
                                #statStateMQTTinternal := #IDLE;
                            END_IF;
                        ELSIF #instTcpSend.ERROR
                        THEN
                            #statusID := #MQTT_PUBLISH;
                            #instTcpSend.REQ := false;
                            #statStateMQTT := #MQTT_ERROR;
                            #status := #instTcpSend.STATUS;
                        END_IF;
                    #MQTT_PUBACK:
                        IF #statNewDataRcv THEN
                            IF ((#statRcvBuffer[1] AND b#16#f0) = #MQTT_MSG_TYPE_PUBACK)
                                OR
                                ((#statRcvBuffer[1] AND b#16#f0) = INT_TO_WORD(#MQTT_MSG_TYPE_PUBREC))
                            THEN
                                IF
                                    (#statRcvBuffer[3] = #statPacketIDAck.%B1)
                                    AND
                                    (#statRcvBuffer[4] = #statPacketIDAck.%B0)
                                THEN
                                    IF (#mqttParam.publishFlag.qualityOfService = 1)
                                    THEN
                                        //QoS = 1; finish here
                                        #statStateMQTTinternal := #MQTT_IDLE;
                                        #published := true;
                                        #busy := false;
                                        #statNewDataRcv := false;
                                        //Re-Activate Kepp Alive Timer
                                        IF NOT #statKeepAliveOff
                                        THEN
                                            #statTriggerKeepAlive := true;
                                        END_IF;

                                        #statStateMQTTinternal := #IDLE;
                                    ELSE
                                        #statStateMQTTinternal := #MQTT_PUBREL;
                                    END_IF;
                                ELSE
                                    #statNewDataRcv := false;
                                END_IF;
                            ELSE
                                #statStateMQTT := #MQTT_ERROR;
                                #statusID := #MQTT_PUBACK;
                            END_IF;
                        END_IF;
                    #MQTT_PUBREL:
                        //fixed Header
                        #statSendBuffer[1] := 16#62;
                        #statSendBuffer[2] := 2;
                        //Variable Header
                        #statSendBuffer[3] := #statPacketID.%B1;
                        #statSendBuffer[4] := #statPacketID.%B0;
                        #instTcpSend.LEN := INT_TO_UDINT(4);
                        #instTcpSend.REQ := true;

                        IF ((#instTcpSend.DONE)
                            AND (#instTcpSend.BUSY = 0))
                        THEN
                            #instTcpSend.REQ := false;
                            #statPacketIDAck := #statPacketID;
                            #statStateMQTTinternal := #MQTT_PUBCOMP;

                        ELSIF #instTcpSend.ERROR
                        THEN
                            #statusID := #MQTT_PUBREL;
                            #instTcpSend.REQ := false;
                            #statStateMQTT := #MQTT_ERROR;
                            #status := #instTcpSend.STATUS;
                        END_IF;
                    #MQTT_PUBCOMP:
                        IF #statNewDataRcv THEN
                            IF ((#statRcvBuffer[1] AND b#16#f0) = #MQTT_MSG_TYPE_PUBCOM)
                            THEN
                                IF
                                    (#statRcvBuffer[3] = #statPacketIDAck.%B1)
                                    AND
                                    (#statRcvBuffer[4] = #statPacketIDAck.%B0)
                                THEN
                                    //QoS = 2; finish here
                                    #statStateMQTTinternal := #MQTT_IDLE;
                                    #published := true;
                                    #busy := false;
                                    #statNewDataRcv := false;
                                    //Re-Activate Kepp Alive Timer
                                    IF NOT #statKeepAliveOff
                                    THEN
                                        #statTriggerKeepAlive := true;
                                    END_IF;

                                    #statStateMQTTinternal := #IDLE;
                                ELSE
                                    #statStateMQTT := #MQTT_ERROR;
                                    #statusID := #MQTT_PUBCOMP;
                                END_IF;
                            END_IF;
                        END_IF;
                    #MQTT_PING:

                        #busy := true;
                        //Build fixed Header
                        //Message Type
                        #statSendBuffer[1] := INT_TO_BYTE(#MQTT_MSG_TYPE_PING);
                        //Remaining Lenght (must be O)
                        #statSendBuffer[2] := 0;
                        #instTcpSend.REQ := true;
                        #instTcpSend.LEN := 2;

                        IF ((#instTcpSend.DONE)
                            AND (#instTcpSend.BUSY = 0))
                        THEN
                            #instTcpSend.REQ := false;
                            #statStateMQTTinternal := #MQTT_PINGRESP;
                        ELSIF #instTcpSend.ERROR
                        THEN
                            #statusID := #MQTT_PING;
                            #instTcpSend.REQ := false;
                            #statStateMQTT := #MQTT_ERROR;
                            #status := #instTcpSend.STATUS;
                        END_IF;
                    #MQTT_PINGRESP:
                        IF #statNewDataRcv
                        THEN
                            IF ((#statRcvBuffer[1] AND b#16#f0) = #MQTT_MSG_TYPE_PINGRESP)
                            THEN
                                #busy := false;
                                #statNewDataRcv := false;
                                #statTriggerKeepAlive := true;
                                #statStateMQTTinternal := #IDLE;
                            END_IF;
                        ELSE
                            #statNewDataRcv := false;
                        END_IF;

                END_CASE;
           #MQTT_DISCONNECT:
           #busy := 0;
           //Build fixed Header
           //Message Type
           #statSendBuffer[1] := INT_TO_BYTE(#MQTT_MSG_TYPE_DISCONNECT);
           //Remaining Lenght (must be O)
           #statSendBuffer[2] := 0;
           #instTcpSend.REQ := true;
           #instTcpSend.LEN := 2;

           IF ((#instTcpSend.DONE)
               AND (#instTcpSend.BUSY = 0))
           THEN
               IF NOT #enable THEN
                   #statStateTCP := #TCP_DISCONNECT;
               END_IF;
               #instTcpSend.REQ := false;
               #statStateMQTT := #MQTT_DISCONNECTED;
               #statStateMQTTinternal := #IDLE;
           ELSIF #instTcpSend.ERROR
           THEN
               IF NOT #enable THEN
                   #statStateTCP := #TCP_DISCONNECT;
               END_IF;
               #statusID := #MQTT_DISCONNECT;
               #instTcpSend.REQ := false;
               #statStateMQTT := #MQTT_ERROR;
               #status := #instTcpSend.STATUS;
           END_IF;
               #MQTT_ERROR:

               REGION Errorhandling MQTT
                   #error := true;
                   #busy := false;
                   #statStateMQTTinternal := #IDLE;
                   #statTriggerKeepAlive := 0;
                   #statKeepAliveOff := false;
                 CASE #statusID OF
                     #MQTT_CONNECT_FLAG_CHECK:
                         #mqttEstablished := false;
                         #statStateMQTT := #MQTT_DISCONNECTED;
                         ;
                     #MQTT_CONNECT:
                         #mqttEstablished := false;
                         #status := #instTcpSend.STATUS;   ;
                         #statStateMQTT := #MQTT_DISCONNECTED;
                       #MQTT_CONNACK:
                           #mqttEstablished := false;
                           #status := #statRcvBuffer[4];
                           #statStateMQTT := #MQTT_DISCONNECTED;
                       #MQTT_PUBLISH:
                               #published := false;
                               #statStateMQTT := #MQTT_CONNECTED;
                               #MQTT_PUBACK,#MQTT_PUBCOMP,#MQTT_PUBREL:
                           #published := false;
                           #status :=#MQTT_ERROR_PACKETID;
                           #statStateMQTT := #MQTT_CONNECTED;
                       #MQTT_PINGRESP:;
                           #MQTT_PING:;
                       #MQTT_DISCONNECT:
                           #mqttEstablished := false;
                          ;
                       ELSE
                           ;
                   END_CASE;
              END_REGION
               ;



       END_CASE
       ;
END_FUNCTION_BLOCK

// folder: NodeRed

FUNCTION "FC_saveMotorDatatoDB" : Void   // FC13, LAD
{ S7_Optimized_Access := 'TRUE' }
VERSION : 0.1
BEGIN

REGION Network 1: M1
   // -temepratura
   // -status POS1
   // -status POS2
   // -isINerror
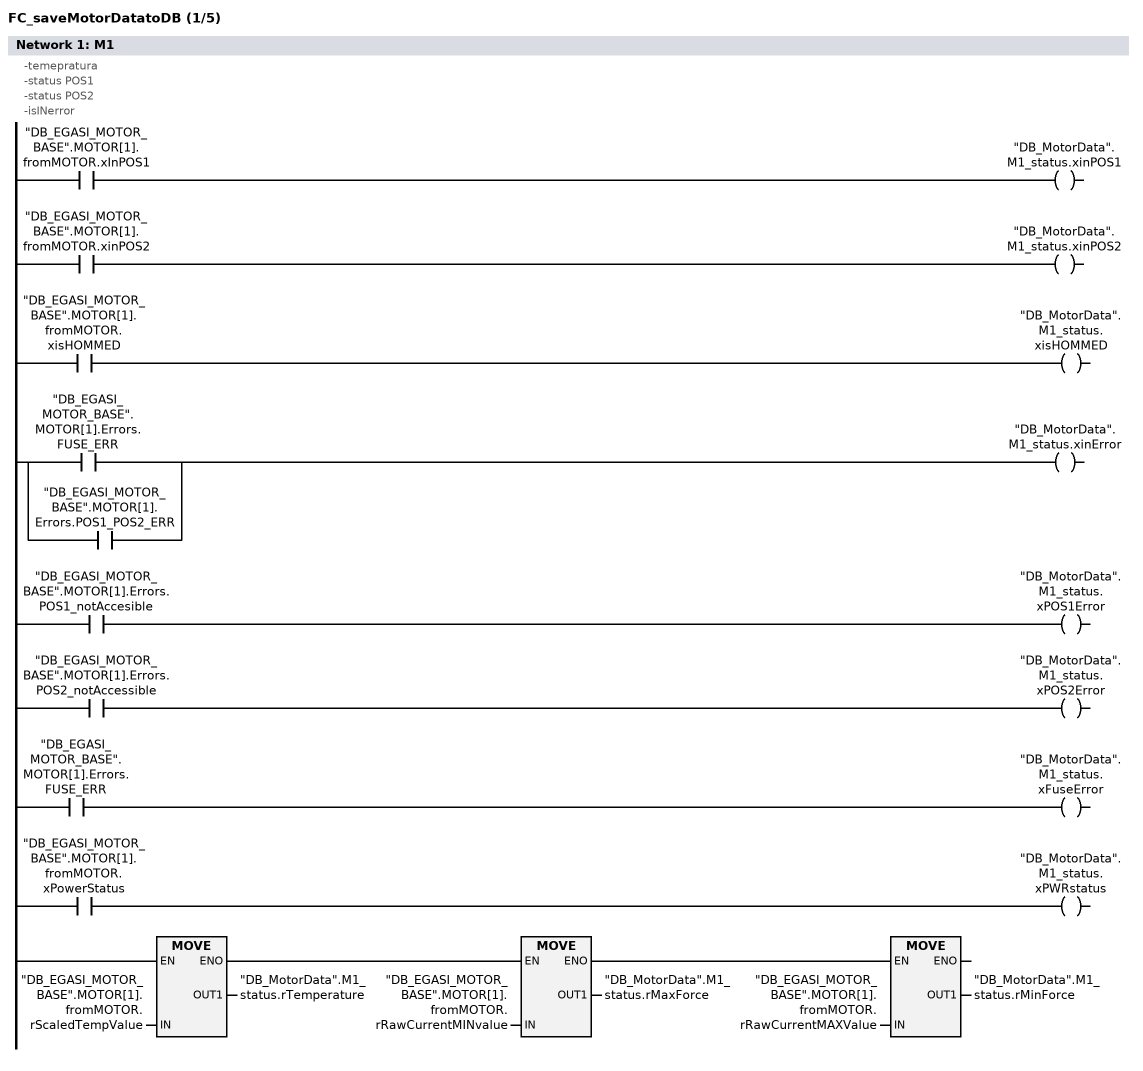
   RUNG wire#powerrail
      Contact( "DB_EGASI_MOTOR_BASE".MOTOR[1].fromMOTOR.xInPOS1 )
      Coil( "DB_MotorData".M1_status.xinPOS1 )
   END_RUNG
   RUNG wire#powerrail
      Contact( "DB_EGASI_MOTOR_BASE".MOTOR[1].fromMOTOR.xinPOS2 )
      Coil( "DB_MotorData".M1_status.xinPOS2 )
   END_RUNG
   RUNG wire#powerrail
      Contact( "DB_EGASI_MOTOR_BASE".MOTOR[1].fromMOTOR.xisHOMMED )
      Coil( "DB_MotorData".M1_status.xisHOMMED )
   END_RUNG
   RUNG wire#powerrail
      Contact( "DB_EGASI_MOTOR_BASE".MOTOR[1].Errors.FUSE_ERR )
      wire#w1
      Coil( "DB_MotorData".M1_status.xinError )
   END_RUNG
   RUNG wire#powerrail
      Contact( "DB_EGASI_MOTOR_BASE".MOTOR[1].Errors.POS1_POS2_ERR )
   END_RUNG wire#w1
   RUNG wire#powerrail
      Contact( "DB_EGASI_MOTOR_BASE".MOTOR[1].Errors.POS1_notAccesible )
      Coil( "DB_MotorData".M1_status.xPOS1Error )
   END_RUNG
   RUNG wire#powerrail
      Contact( "DB_EGASI_MOTOR_BASE".MOTOR[1].Errors.POS2_notAccessible )
      Coil( "DB_MotorData".M1_status.xPOS2Error )
   END_RUNG
   RUNG wire#powerrail
      Contact( "DB_EGASI_MOTOR_BASE".MOTOR[1].Errors.FUSE_ERR )
      Coil( "DB_MotorData".M1_status.xFuseError )
   END_RUNG
   RUNG wire#powerrail
      Contact( "DB_EGASI_MOTOR_BASE".MOTOR[1].fromMOTOR.xPowerStatus )
      Coil( "DB_MotorData".M1_status.xPWRstatus )
   END_RUNG
   RUNG wire#powerrail
      Move(in := "DB_EGASI_MOTOR_BASE".MOTOR[1].fromMOTOR.rScaledTempValue, out1 => "DB_MotorData".M1_status.rTemperature)
      Move(in := "DB_EGASI_MOTOR_BASE".MOTOR[1].fromMOTOR.rRawCurrentMINvalue, out1 => "DB_MotorData".M1_status.rMaxForce)
      Move(in := "DB_EGASI_MOTOR_BASE".MOTOR[1].fromMOTOR.rRawCurrentMAXValue, out1 => "DB_MotorData".M1_status.rMinForce)
   END_RUNG
   // the same network as SCL:
   "DB_MotorData".M1_status.xinPOS1 := "DB_EGASI_MOTOR_BASE".MOTOR[1].fromMOTOR.xInPOS1;
   "DB_MotorData".M1_status.xinPOS2 := "DB_EGASI_MOTOR_BASE".MOTOR[1].fromMOTOR.xinPOS2;
   "DB_MotorData".M1_status.xisHOMMED := "DB_EGASI_MOTOR_BASE".MOTOR[1].fromMOTOR.xisHOMMED;
   "DB_MotorData".M1_status.xinError := "DB_EGASI_MOTOR_BASE".MOTOR[1].Errors.FUSE_ERR OR "DB_EGASI_MOTOR_BASE".MOTOR[1].Errors.POS1_POS2_ERR;
   "DB_MotorData".M1_status.xPOS1Error := "DB_EGASI_MOTOR_BASE".MOTOR[1].Errors.POS1_notAccesible;
   "DB_MotorData".M1_status.xPOS2Error := "DB_EGASI_MOTOR_BASE".MOTOR[1].Errors.POS2_notAccessible;
   "DB_MotorData".M1_status.xFuseError := "DB_EGASI_MOTOR_BASE".MOTOR[1].Errors.FUSE_ERR;
   "DB_MotorData".M1_status.xPWRstatus := "DB_EGASI_MOTOR_BASE".MOTOR[1].fromMOTOR.xPowerStatus;
   "DB_MotorData".M1_status.rTemperature := "DB_EGASI_MOTOR_BASE".MOTOR[1].fromMOTOR.rScaledTempValue;
   "DB_MotorData".M1_status.rMaxForce := "DB_EGASI_MOTOR_BASE".MOTOR[1].fromMOTOR.rRawCurrentMINvalue;
   "DB_MotorData".M1_status.rMinForce := "DB_EGASI_MOTOR_BASE".MOTOR[1].fromMOTOR.rRawCurrentMAXValue;
END_REGION

REGION Network 2: M2
   // -temepratura
   // -status POS1
   // -status POS2
   // -isINerror
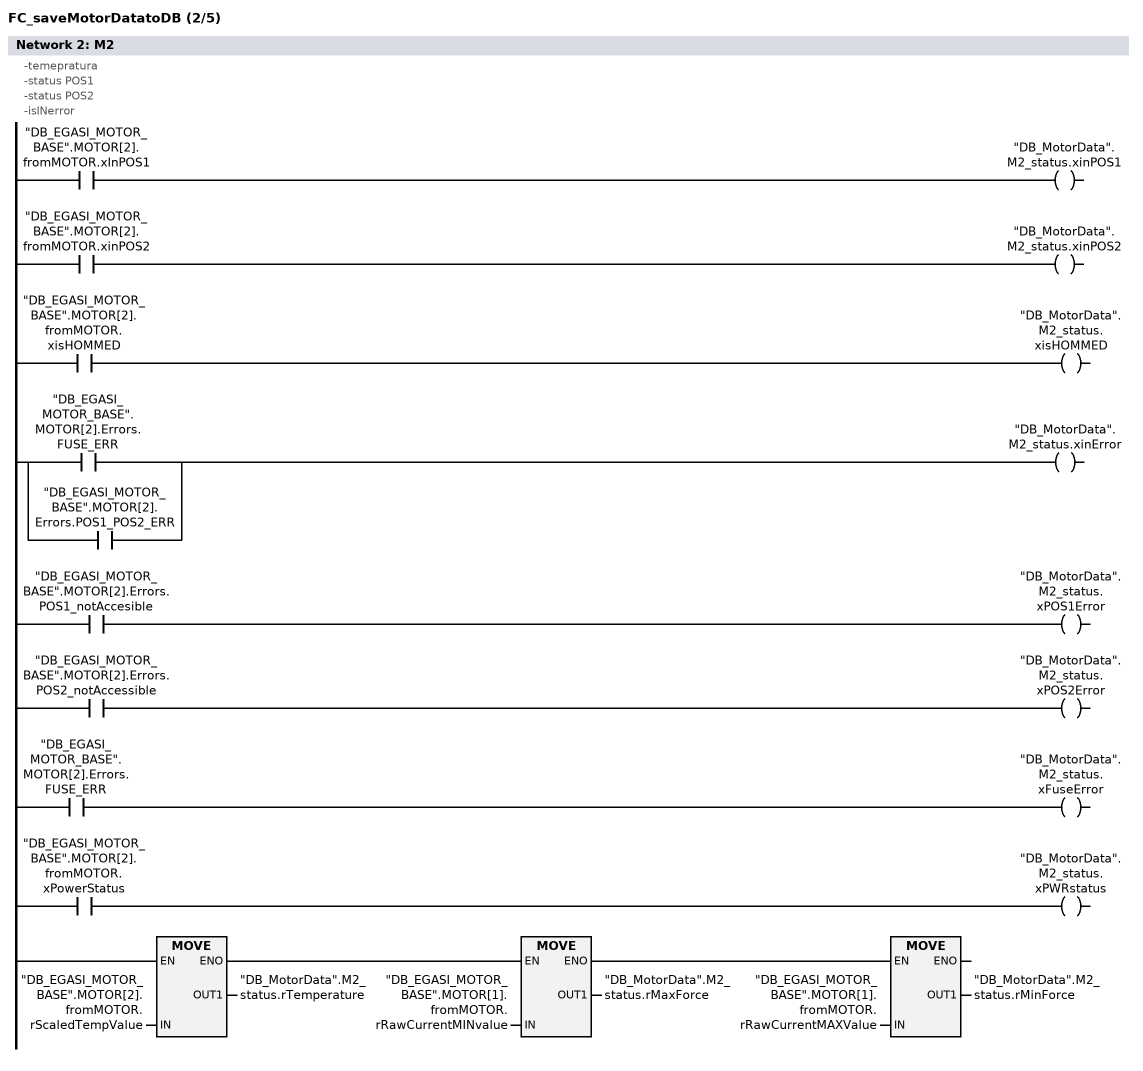
   RUNG wire#powerrail
      Contact( "DB_EGASI_MOTOR_BASE".MOTOR[2].fromMOTOR.xInPOS1 )
      Coil( "DB_MotorData".M2_status.xinPOS1 )
   END_RUNG
   RUNG wire#powerrail
      Contact( "DB_EGASI_MOTOR_BASE".MOTOR[2].fromMOTOR.xinPOS2 )
      Coil( "DB_MotorData".M2_status.xinPOS2 )
   END_RUNG
   RUNG wire#powerrail
      Contact( "DB_EGASI_MOTOR_BASE".MOTOR[2].fromMOTOR.xisHOMMED )
      Coil( "DB_MotorData".M2_status.xisHOMMED )
   END_RUNG
   RUNG wire#powerrail
      Contact( "DB_EGASI_MOTOR_BASE".MOTOR[2].Errors.FUSE_ERR )
      wire#w1
      Coil( "DB_MotorData".M2_status.xinError )
   END_RUNG
   RUNG wire#powerrail
      Contact( "DB_EGASI_MOTOR_BASE".MOTOR[2].Errors.POS1_POS2_ERR )
   END_RUNG wire#w1
   RUNG wire#powerrail
      Contact( "DB_EGASI_MOTOR_BASE".MOTOR[2].Errors.POS1_notAccesible )
      Coil( "DB_MotorData".M2_status.xPOS1Error )
   END_RUNG
   RUNG wire#powerrail
      Contact( "DB_EGASI_MOTOR_BASE".MOTOR[2].Errors.POS2_notAccessible )
      Coil( "DB_MotorData".M2_status.xPOS2Error )
   END_RUNG
   RUNG wire#powerrail
      Contact( "DB_EGASI_MOTOR_BASE".MOTOR[2].Errors.FUSE_ERR )
      Coil( "DB_MotorData".M2_status.xFuseError )
   END_RUNG
   RUNG wire#powerrail
      Contact( "DB_EGASI_MOTOR_BASE".MOTOR[2].fromMOTOR.xPowerStatus )
      Coil( "DB_MotorData".M2_status.xPWRstatus )
   END_RUNG
   RUNG wire#powerrail
      Move(in := "DB_EGASI_MOTOR_BASE".MOTOR[2].fromMOTOR.rScaledTempValue, out1 => "DB_MotorData".M2_status.rTemperature)
      Move(in := "DB_EGASI_MOTOR_BASE".MOTOR[1].fromMOTOR.rRawCurrentMINvalue, out1 => "DB_MotorData".M2_status.rMaxForce)
      Move(in := "DB_EGASI_MOTOR_BASE".MOTOR[1].fromMOTOR.rRawCurrentMAXValue, out1 => "DB_MotorData".M2_status.rMinForce)
   END_RUNG
   // the same network as SCL:
   "DB_MotorData".M2_status.xinPOS1 := "DB_EGASI_MOTOR_BASE".MOTOR[2].fromMOTOR.xInPOS1;
   "DB_MotorData".M2_status.xinPOS2 := "DB_EGASI_MOTOR_BASE".MOTOR[2].fromMOTOR.xinPOS2;
   "DB_MotorData".M2_status.xisHOMMED := "DB_EGASI_MOTOR_BASE".MOTOR[2].fromMOTOR.xisHOMMED;
   "DB_MotorData".M2_status.xinError := "DB_EGASI_MOTOR_BASE".MOTOR[2].Errors.FUSE_ERR OR "DB_EGASI_MOTOR_BASE".MOTOR[2].Errors.POS1_POS2_ERR;
   "DB_MotorData".M2_status.xPOS1Error := "DB_EGASI_MOTOR_BASE".MOTOR[2].Errors.POS1_notAccesible;
   "DB_MotorData".M2_status.xPOS2Error := "DB_EGASI_MOTOR_BASE".MOTOR[2].Errors.POS2_notAccessible;
   "DB_MotorData".M2_status.xFuseError := "DB_EGASI_MOTOR_BASE".MOTOR[2].Errors.FUSE_ERR;
   "DB_MotorData".M2_status.xPWRstatus := "DB_EGASI_MOTOR_BASE".MOTOR[2].fromMOTOR.xPowerStatus;
   "DB_MotorData".M2_status.rTemperature := "DB_EGASI_MOTOR_BASE".MOTOR[2].fromMOTOR.rScaledTempValue;
   "DB_MotorData".M2_status.rMaxForce := "DB_EGASI_MOTOR_BASE".MOTOR[1].fromMOTOR.rRawCurrentMINvalue;
   "DB_MotorData".M2_status.rMinForce := "DB_EGASI_MOTOR_BASE".MOTOR[1].fromMOTOR.rRawCurrentMAXValue;
END_REGION

REGION Network 3: M3
   // -temepratura
   // -status POS1
   // -status POS2
   // -isINerror
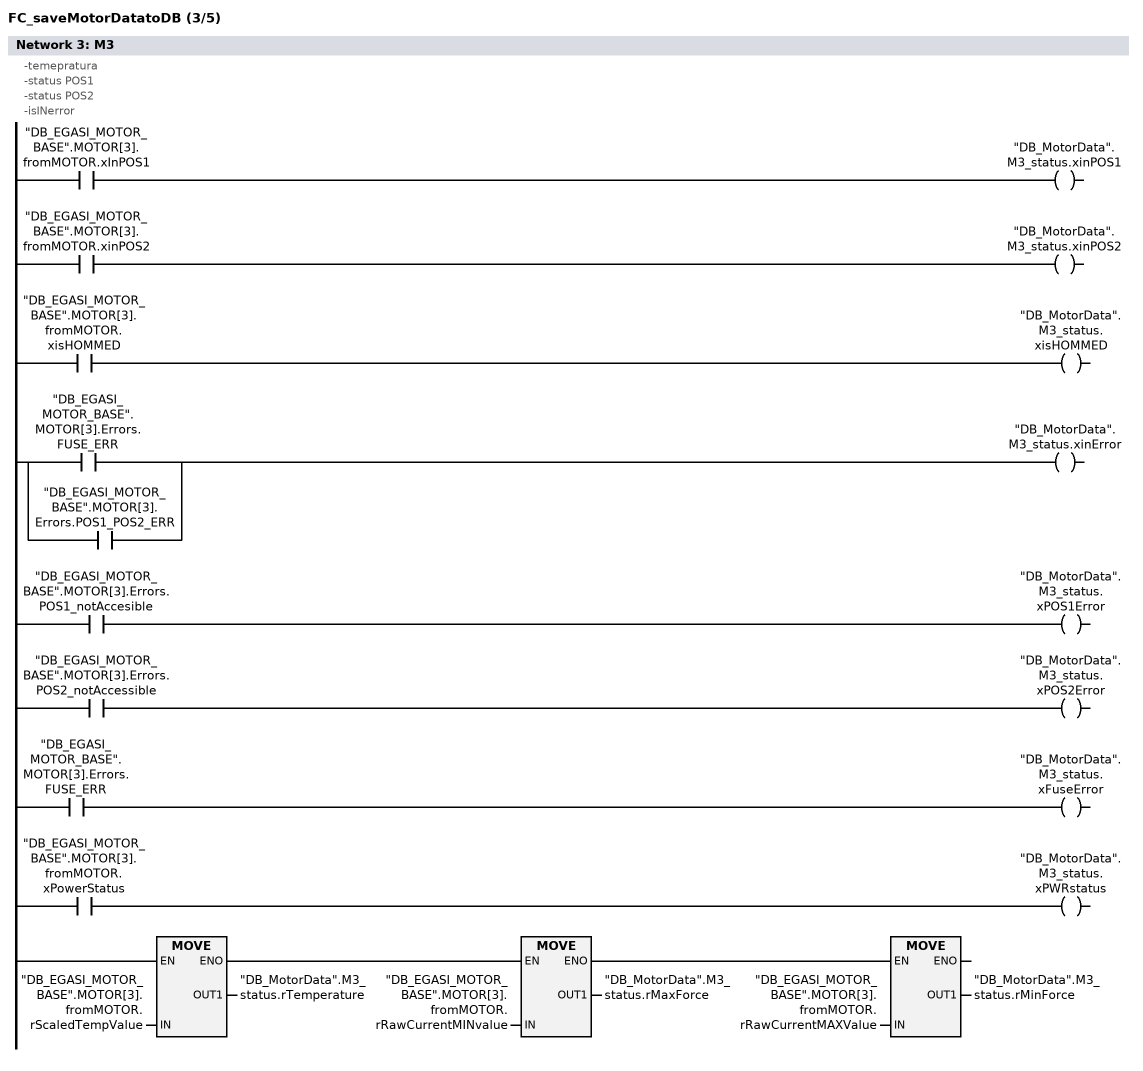
   RUNG wire#powerrail
      Contact( "DB_EGASI_MOTOR_BASE".MOTOR[3].fromMOTOR.xInPOS1 )
      Coil( "DB_MotorData".M3_status.xinPOS1 )
   END_RUNG
   RUNG wire#powerrail
      Contact( "DB_EGASI_MOTOR_BASE".MOTOR[3].fromMOTOR.xinPOS2 )
      Coil( "DB_MotorData".M3_status.xinPOS2 )
   END_RUNG
   RUNG wire#powerrail
      Contact( "DB_EGASI_MOTOR_BASE".MOTOR[3].fromMOTOR.xisHOMMED )
      Coil( "DB_MotorData".M3_status.xisHOMMED )
   END_RUNG
   RUNG wire#powerrail
      Contact( "DB_EGASI_MOTOR_BASE".MOTOR[3].Errors.FUSE_ERR )
      wire#w1
      Coil( "DB_MotorData".M3_status.xinError )
   END_RUNG
   RUNG wire#powerrail
      Contact( "DB_EGASI_MOTOR_BASE".MOTOR[3].Errors.POS1_POS2_ERR )
   END_RUNG wire#w1
   RUNG wire#powerrail
      Contact( "DB_EGASI_MOTOR_BASE".MOTOR[3].Errors.POS1_notAccesible )
      Coil( "DB_MotorData".M3_status.xPOS1Error )
   END_RUNG
   RUNG wire#powerrail
      Contact( "DB_EGASI_MOTOR_BASE".MOTOR[3].Errors.POS2_notAccessible )
      Coil( "DB_MotorData".M3_status.xPOS2Error )
   END_RUNG
   RUNG wire#powerrail
      Contact( "DB_EGASI_MOTOR_BASE".MOTOR[3].Errors.FUSE_ERR )
      Coil( "DB_MotorData".M3_status.xFuseError )
   END_RUNG
   RUNG wire#powerrail
      Contact( "DB_EGASI_MOTOR_BASE".MOTOR[3].fromMOTOR.xPowerStatus )
      Coil( "DB_MotorData".M3_status.xPWRstatus )
   END_RUNG
   RUNG wire#powerrail
      Move(in := "DB_EGASI_MOTOR_BASE".MOTOR[3].fromMOTOR.rScaledTempValue, out1 => "DB_MotorData".M3_status.rTemperature)
      Move(in := "DB_EGASI_MOTOR_BASE".MOTOR[3].fromMOTOR.rRawCurrentMINvalue, out1 => "DB_MotorData".M3_status.rMaxForce)
      Move(in := "DB_EGASI_MOTOR_BASE".MOTOR[3].fromMOTOR.rRawCurrentMAXValue, out1 => "DB_MotorData".M3_status.rMinForce)
   END_RUNG
   // the same network as SCL:
   "DB_MotorData".M3_status.xinPOS1 := "DB_EGASI_MOTOR_BASE".MOTOR[3].fromMOTOR.xInPOS1;
   "DB_MotorData".M3_status.xinPOS2 := "DB_EGASI_MOTOR_BASE".MOTOR[3].fromMOTOR.xinPOS2;
   "DB_MotorData".M3_status.xisHOMMED := "DB_EGASI_MOTOR_BASE".MOTOR[3].fromMOTOR.xisHOMMED;
   "DB_MotorData".M3_status.xinError := "DB_EGASI_MOTOR_BASE".MOTOR[3].Errors.FUSE_ERR OR "DB_EGASI_MOTOR_BASE".MOTOR[3].Errors.POS1_POS2_ERR;
   "DB_MotorData".M3_status.xPOS1Error := "DB_EGASI_MOTOR_BASE".MOTOR[3].Errors.POS1_notAccesible;
   "DB_MotorData".M3_status.xPOS2Error := "DB_EGASI_MOTOR_BASE".MOTOR[3].Errors.POS2_notAccessible;
   "DB_MotorData".M3_status.xFuseError := "DB_EGASI_MOTOR_BASE".MOTOR[3].Errors.FUSE_ERR;
   "DB_MotorData".M3_status.xPWRstatus := "DB_EGASI_MOTOR_BASE".MOTOR[3].fromMOTOR.xPowerStatus;
   "DB_MotorData".M3_status.rTemperature := "DB_EGASI_MOTOR_BASE".MOTOR[3].fromMOTOR.rScaledTempValue;
   "DB_MotorData".M3_status.rMaxForce := "DB_EGASI_MOTOR_BASE".MOTOR[3].fromMOTOR.rRawCurrentMINvalue;
   "DB_MotorData".M3_status.rMinForce := "DB_EGASI_MOTOR_BASE".MOTOR[3].fromMOTOR.rRawCurrentMAXValue;
END_REGION

REGION Network 4: M4
   // -temepratura
   // -status POS1
   // -status POS2
   // -isINerror
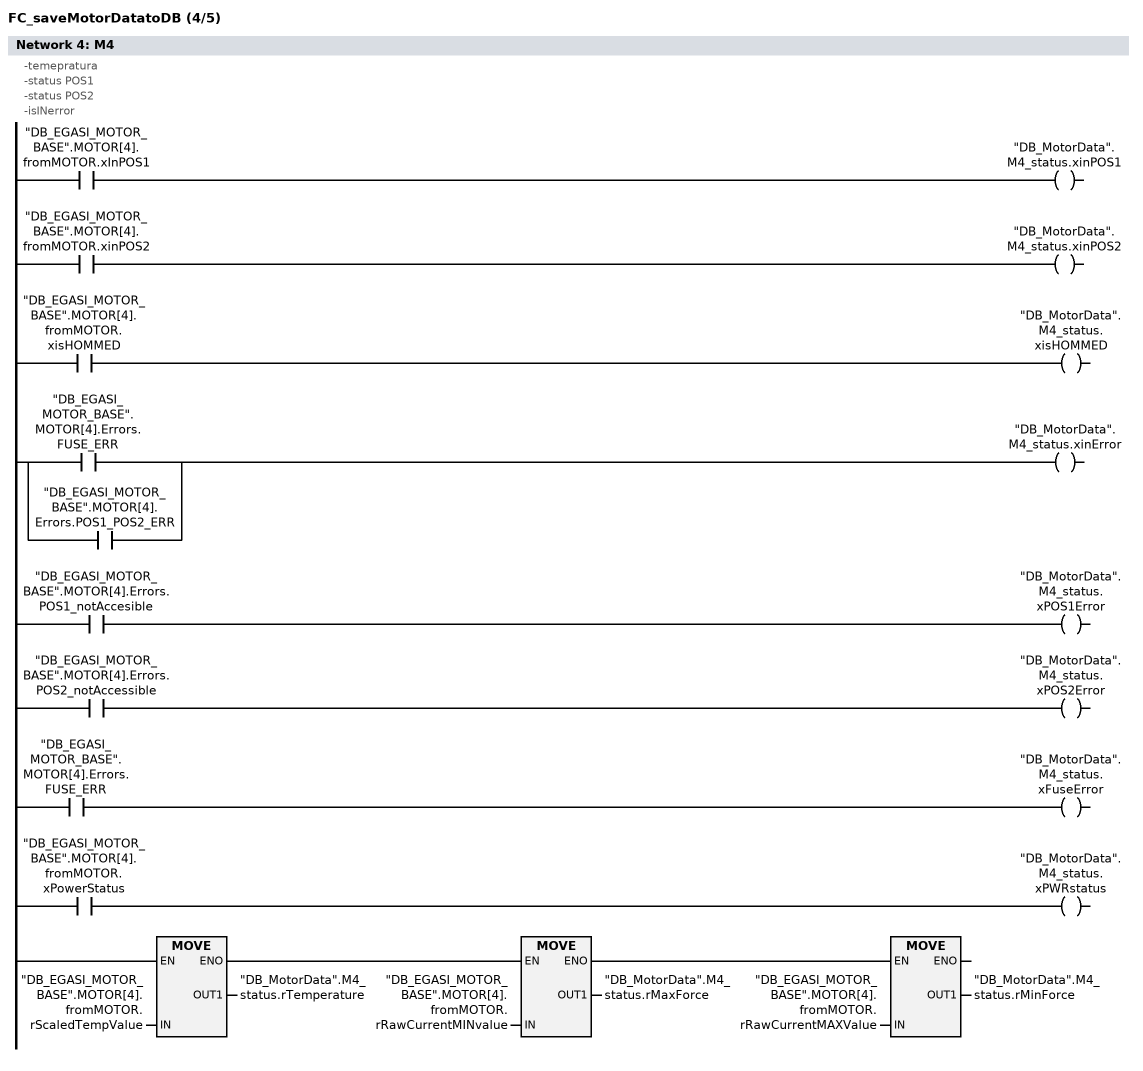
   RUNG wire#powerrail
      Contact( "DB_EGASI_MOTOR_BASE".MOTOR[4].fromMOTOR.xInPOS1 )
      Coil( "DB_MotorData".M4_status.xinPOS1 )
   END_RUNG
   RUNG wire#powerrail
      Contact( "DB_EGASI_MOTOR_BASE".MOTOR[4].fromMOTOR.xinPOS2 )
      Coil( "DB_MotorData".M4_status.xinPOS2 )
   END_RUNG
   RUNG wire#powerrail
      Contact( "DB_EGASI_MOTOR_BASE".MOTOR[4].fromMOTOR.xisHOMMED )
      Coil( "DB_MotorData".M4_status.xisHOMMED )
   END_RUNG
   RUNG wire#powerrail
      Contact( "DB_EGASI_MOTOR_BASE".MOTOR[4].Errors.FUSE_ERR )
      wire#w1
      Coil( "DB_MotorData".M4_status.xinError )
   END_RUNG
   RUNG wire#powerrail
      Contact( "DB_EGASI_MOTOR_BASE".MOTOR[4].Errors.POS1_POS2_ERR )
   END_RUNG wire#w1
   RUNG wire#powerrail
      Contact( "DB_EGASI_MOTOR_BASE".MOTOR[4].Errors.POS1_notAccesible )
      Coil( "DB_MotorData".M4_status.xPOS1Error )
   END_RUNG
   RUNG wire#powerrail
      Contact( "DB_EGASI_MOTOR_BASE".MOTOR[4].Errors.POS2_notAccessible )
      Coil( "DB_MotorData".M4_status.xPOS2Error )
   END_RUNG
   RUNG wire#powerrail
      Contact( "DB_EGASI_MOTOR_BASE".MOTOR[4].Errors.FUSE_ERR )
      Coil( "DB_MotorData".M4_status.xFuseError )
   END_RUNG
   RUNG wire#powerrail
      Contact( "DB_EGASI_MOTOR_BASE".MOTOR[4].fromMOTOR.xPowerStatus )
      Coil( "DB_MotorData".M4_status.xPWRstatus )
   END_RUNG
   RUNG wire#powerrail
      Move(in := "DB_EGASI_MOTOR_BASE".MOTOR[4].fromMOTOR.rScaledTempValue, out1 => "DB_MotorData".M4_status.rTemperature)
      Move(in := "DB_EGASI_MOTOR_BASE".MOTOR[4].fromMOTOR.rRawCurrentMINvalue, out1 => "DB_MotorData".M4_status.rMaxForce)
      Move(in := "DB_EGASI_MOTOR_BASE".MOTOR[4].fromMOTOR.rRawCurrentMAXValue, out1 => "DB_MotorData".M4_status.rMinForce)
   END_RUNG
   // the same network as SCL:
   "DB_MotorData".M4_status.xinPOS1 := "DB_EGASI_MOTOR_BASE".MOTOR[4].fromMOTOR.xInPOS1;
   "DB_MotorData".M4_status.xinPOS2 := "DB_EGASI_MOTOR_BASE".MOTOR[4].fromMOTOR.xinPOS2;
   "DB_MotorData".M4_status.xisHOMMED := "DB_EGASI_MOTOR_BASE".MOTOR[4].fromMOTOR.xisHOMMED;
   "DB_MotorData".M4_status.xinError := "DB_EGASI_MOTOR_BASE".MOTOR[4].Errors.FUSE_ERR OR "DB_EGASI_MOTOR_BASE".MOTOR[4].Errors.POS1_POS2_ERR;
   "DB_MotorData".M4_status.xPOS1Error := "DB_EGASI_MOTOR_BASE".MOTOR[4].Errors.POS1_notAccesible;
   "DB_MotorData".M4_status.xPOS2Error := "DB_EGASI_MOTOR_BASE".MOTOR[4].Errors.POS2_notAccessible;
   "DB_MotorData".M4_status.xFuseError := "DB_EGASI_MOTOR_BASE".MOTOR[4].Errors.FUSE_ERR;
   "DB_MotorData".M4_status.xPWRstatus := "DB_EGASI_MOTOR_BASE".MOTOR[4].fromMOTOR.xPowerStatus;
   "DB_MotorData".M4_status.rTemperature := "DB_EGASI_MOTOR_BASE".MOTOR[4].fromMOTOR.rScaledTempValue;
   "DB_MotorData".M4_status.rMaxForce := "DB_EGASI_MOTOR_BASE".MOTOR[4].fromMOTOR.rRawCurrentMINvalue;
   "DB_MotorData".M4_status.rMinForce := "DB_EGASI_MOTOR_BASE".MOTOR[4].fromMOTOR.rRawCurrentMAXValue;
END_REGION

REGION Network 5: M5
   // -temepratura
   // -status POS1
   // -status POS2
   // -isINerror
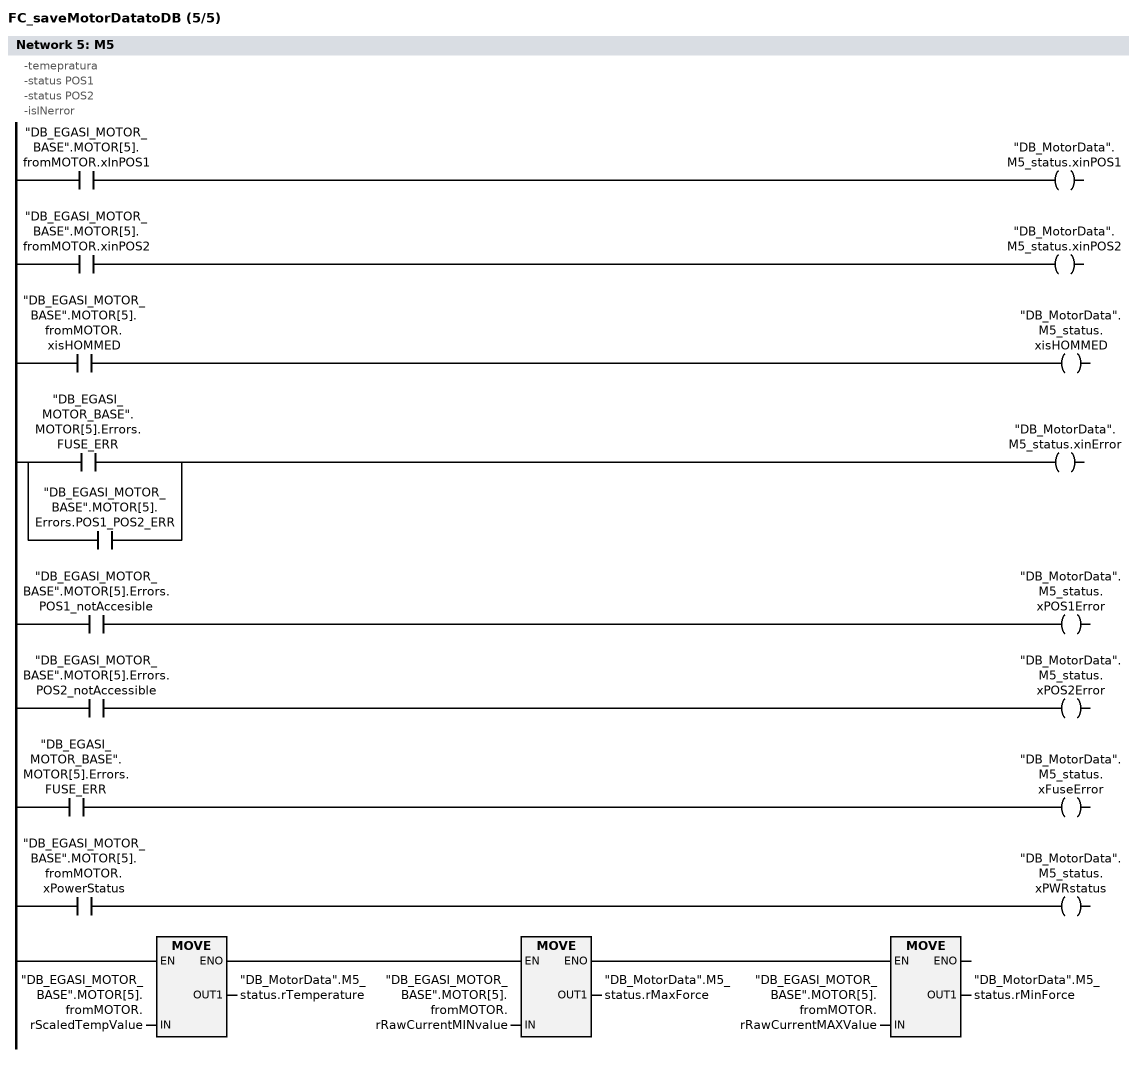
   RUNG wire#powerrail
      Contact( "DB_EGASI_MOTOR_BASE".MOTOR[5].fromMOTOR.xInPOS1 )
      Coil( "DB_MotorData".M5_status.xinPOS1 )
   END_RUNG
   RUNG wire#powerrail
      Contact( "DB_EGASI_MOTOR_BASE".MOTOR[5].fromMOTOR.xinPOS2 )
      Coil( "DB_MotorData".M5_status.xinPOS2 )
   END_RUNG
   RUNG wire#powerrail
      Contact( "DB_EGASI_MOTOR_BASE".MOTOR[5].fromMOTOR.xisHOMMED )
      Coil( "DB_MotorData".M5_status.xisHOMMED )
   END_RUNG
   RUNG wire#powerrail
      Contact( "DB_EGASI_MOTOR_BASE".MOTOR[5].Errors.FUSE_ERR )
      wire#w1
      Coil( "DB_MotorData".M5_status.xinError )
   END_RUNG
   RUNG wire#powerrail
      Contact( "DB_EGASI_MOTOR_BASE".MOTOR[5].Errors.POS1_POS2_ERR )
   END_RUNG wire#w1
   RUNG wire#powerrail
      Contact( "DB_EGASI_MOTOR_BASE".MOTOR[5].Errors.POS1_notAccesible )
      Coil( "DB_MotorData".M5_status.xPOS1Error )
   END_RUNG
   RUNG wire#powerrail
      Contact( "DB_EGASI_MOTOR_BASE".MOTOR[5].Errors.POS2_notAccessible )
      Coil( "DB_MotorData".M5_status.xPOS2Error )
   END_RUNG
   RUNG wire#powerrail
      Contact( "DB_EGASI_MOTOR_BASE".MOTOR[5].Errors.FUSE_ERR )
      Coil( "DB_MotorData".M5_status.xFuseError )
   END_RUNG
   RUNG wire#powerrail
      Contact( "DB_EGASI_MOTOR_BASE".MOTOR[5].fromMOTOR.xPowerStatus )
      Coil( "DB_MotorData".M5_status.xPWRstatus )
   END_RUNG
   RUNG wire#powerrail
      Move(in := "DB_EGASI_MOTOR_BASE".MOTOR[5].fromMOTOR.rScaledTempValue, out1 => "DB_MotorData".M5_status.rTemperature)
      Move(in := "DB_EGASI_MOTOR_BASE".MOTOR[5].fromMOTOR.rRawCurrentMINvalue, out1 => "DB_MotorData".M5_status.rMaxForce)
      Move(in := "DB_EGASI_MOTOR_BASE".MOTOR[5].fromMOTOR.rRawCurrentMAXValue, out1 => "DB_MotorData".M5_status.rMinForce)
   END_RUNG
   // the same network as SCL:
   "DB_MotorData".M5_status.xinPOS1 := "DB_EGASI_MOTOR_BASE".MOTOR[5].fromMOTOR.xInPOS1;
   "DB_MotorData".M5_status.xinPOS2 := "DB_EGASI_MOTOR_BASE".MOTOR[5].fromMOTOR.xinPOS2;
   "DB_MotorData".M5_status.xisHOMMED := "DB_EGASI_MOTOR_BASE".MOTOR[5].fromMOTOR.xisHOMMED;
   "DB_MotorData".M5_status.xinError := "DB_EGASI_MOTOR_BASE".MOTOR[5].Errors.FUSE_ERR OR "DB_EGASI_MOTOR_BASE".MOTOR[5].Errors.POS1_POS2_ERR;
   "DB_MotorData".M5_status.xPOS1Error := "DB_EGASI_MOTOR_BASE".MOTOR[5].Errors.POS1_notAccesible;
   "DB_MotorData".M5_status.xPOS2Error := "DB_EGASI_MOTOR_BASE".MOTOR[5].Errors.POS2_notAccessible;
   "DB_MotorData".M5_status.xFuseError := "DB_EGASI_MOTOR_BASE".MOTOR[5].Errors.FUSE_ERR;
   "DB_MotorData".M5_status.xPWRstatus := "DB_EGASI_MOTOR_BASE".MOTOR[5].fromMOTOR.xPowerStatus;
   "DB_MotorData".M5_status.rTemperature := "DB_EGASI_MOTOR_BASE".MOTOR[5].fromMOTOR.rScaledTempValue;
   "DB_MotorData".M5_status.rMaxForce := "DB_EGASI_MOTOR_BASE".MOTOR[5].fromMOTOR.rRawCurrentMINvalue;
   "DB_MotorData".M5_status.rMinForce := "DB_EGASI_MOTOR_BASE".MOTOR[5].fromMOTOR.rRawCurrentMAXValue;
END_REGION
END_FUNCTION